// TIA Portal project "Inteligenta_szklarnia" (V15.1) (continued)
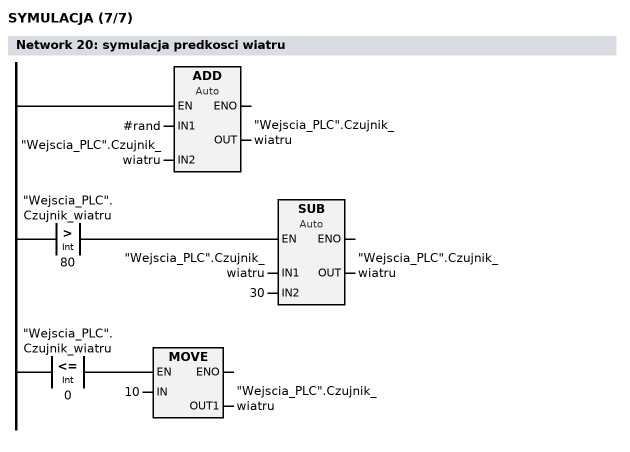
   RUNG wire#powerrail
      Add(in1 := #rand, in2 := "Wejscia_PLC".Czujnik_wiatru, out => "Wejscia_PLC".Czujnik_wiatru)
   END_RUNG
   RUNG wire#powerrail
      { S7_Templates := "SrcType := Int" } GT_Contact(in1 := "Wejscia_PLC".Czujnik_wiatru, in2 := 80)
      Sub(in1 := "Wejscia_PLC".Czujnik_wiatru, in2 := 30, out => "Wejscia_PLC".Czujnik_wiatru)
   END_RUNG
   RUNG wire#powerrail
      { S7_Templates := "SrcType := Int" } LE_Contact(in1 := "Wejscia_PLC".Czujnik_wiatru, in2 := 0)
      Move(in := 10, out1 => "Wejscia_PLC".Czujnik_wiatru)
   END_RUNG
   // the same network as SCL:
   "Wejscia_PLC".Czujnik_wiatru := #rand + "Wejscia_PLC".Czujnik_wiatru;
   IF "Wejscia_PLC".Czujnik_wiatru > 80 THEN
       "Wejscia_PLC".Czujnik_wiatru := "Wejscia_PLC".Czujnik_wiatru - 30;
   END_IF;
   IF "Wejscia_PLC".Czujnik_wiatru <= 0 THEN "Wejscia_PLC".Czujnik_wiatru := 10; END_IF;
END_REGION
END_FUNCTION

ORGANIZATION_BLOCK "Main"   // OB1, LAD, ProgramCycle
TITLE = "Main Program Sweep (Cycle)"
{ S7_Optimized_Access := 'TRUE' }
VERSION : 0.1
   VAR_INPUT
      Initial_Call : Bool;   // Initial call of this OB
      Remanence : Bool;   // =True, if remanent data are available
   END_VAR
   VAR_TEMP   // added for the SCL form of the ladder/FBD networks
      _w1 : Bool;
   END_VAR
BEGIN

REGION Network 1
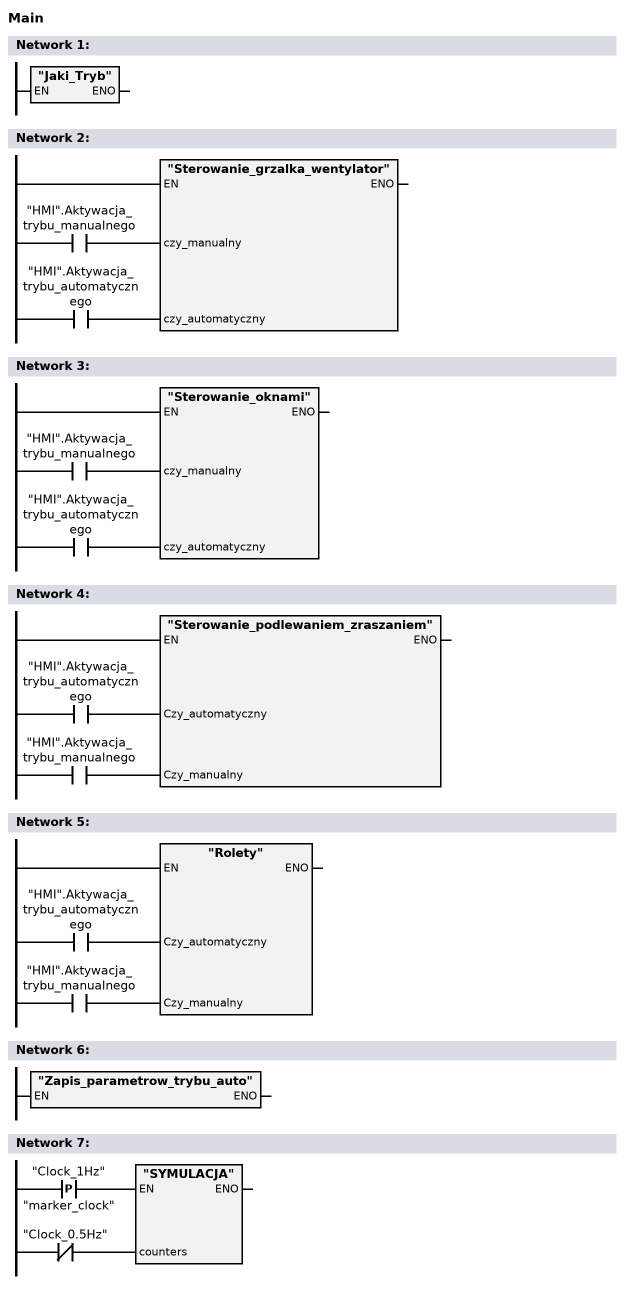
   RUNG wire#powerrail
      "Jaki_Tryb"()
   END_RUNG
   // the same network as SCL:
   "Jaki_Tryb"();
END_REGION

REGION Network 2
   RUNG wire#powerrail
      "Sterowanie_grzalka_wentylator"(czy_manualny := wire#w1, czy_automatyczny := wire#w2)
   END_RUNG
   RUNG wire#powerrail
      Contact( "HMI".Aktywacja_trybu_manualnego )
   END_RUNG wire#w1
   RUNG wire#powerrail
      Contact( "HMI".Aktywacja_trybu_automatycznego )
   END_RUNG wire#w2
   // the same network as SCL:
   "Sterowanie_grzalka_wentylator"(czy_manualny := "HMI".Aktywacja_trybu_manualnego,
                           czy_automatyczny := "HMI".Aktywacja_trybu_automatycznego);
END_REGION

REGION Network 3
   RUNG wire#powerrail
      "Sterowanie_oknami"(czy_manualny := wire#w1, czy_automatyczny := wire#w2)
   END_RUNG
   RUNG wire#powerrail
      Contact( "HMI".Aktywacja_trybu_manualnego )
   END_RUNG wire#w1
   RUNG wire#powerrail
      Contact( "HMI".Aktywacja_trybu_automatycznego )
   END_RUNG wire#w2
   // the same network as SCL:
   "Sterowanie_oknami"(czy_manualny := "HMI".Aktywacja_trybu_manualnego,
                       czy_automatyczny := "HMI".Aktywacja_trybu_automatycznego);
END_REGION

REGION Network 4
   RUNG wire#powerrail
      "Sterowanie_podlewaniem_zraszaniem"(Czy_automatyczny := wire#w1, Czy_manualny := wire#w2)
   END_RUNG
   RUNG wire#powerrail
      Contact( "HMI".Aktywacja_trybu_automatycznego )
   END_RUNG wire#w1
   RUNG wire#powerrail
      Contact( "HMI".Aktywacja_trybu_manualnego )
   END_RUNG wire#w2
   // the same network as SCL:
   "Sterowanie_podlewaniem_zraszaniem"(Czy_automatyczny := "HMI".Aktywacja_trybu_automatycznego,
                           Czy_manualny := "HMI".Aktywacja_trybu_manualnego);
END_REGION

REGION Network 5
   RUNG wire#powerrail
      "Rolety"(Czy_automatyczny := wire#w1, Czy_manualny := wire#w2)
   END_RUNG
   RUNG wire#powerrail
      Contact( "HMI".Aktywacja_trybu_automatycznego )
   END_RUNG wire#w1
   RUNG wire#powerrail
      Contact( "HMI".Aktywacja_trybu_manualnego )
   END_RUNG wire#w2
   // the same network as SCL:
   "Rolety"(Czy_automatyczny := "HMI".Aktywacja_trybu_automatycznego,
            Czy_manualny := "HMI".Aktywacja_trybu_manualnego);
END_REGION

REGION Network 6
   RUNG wire#powerrail
      "Zapis_parametrow_trybu_auto"()
   END_RUNG
   // the same network as SCL:
   "Zapis_parametrow_trybu_auto"();
END_REGION

REGION Network 7
   RUNG wire#powerrail
      P_Contact(operand := "Clock_1Hz", bit := "marker_clock")
      "SYMULACJA"(counters := wire#w1)
   END_RUNG
   RUNG wire#powerrail
      I_Contact( "Clock_0.5Hz" )
   END_RUNG wire#w1
   // the same network as SCL:
   #_w1 := "Clock_1Hz" AND NOT "marker_clock";   // rising edge of "Clock_1Hz"
   "marker_clock" := "Clock_1Hz";
   IF #_w1 THEN "SYMULACJA"(counters := NOT "Clock_0.5Hz"); END_IF;
END_REGION
END_ORGANIZATION_BLOCK

// folder: Archiwizacja_parametrow

FUNCTION "Archiwizacja_parametrow" : Void   // FC2, LAD
{ S7_Optimized_Access := 'TRUE' }
VERSION : 0.1
// Zapis parametrów do bloku DB odbywa się co pół godziny. Po uruchomieniu sterownika pierwszy zapis nie odbywa się od razu, aby wykres nie przedstawiał parametrów, które nie były jeszcze regulowane. Oczytane watosci zapisywane są w tablicach w bloku DB.
   VAR CONSTANT
      iterator : Int := 0;
   END_VAR
   VAR_TEMP   // added for the SCL form of the ladder/FBD networks
      _w1 : Bool;
   END_VAR
BEGIN

REGION Network 1
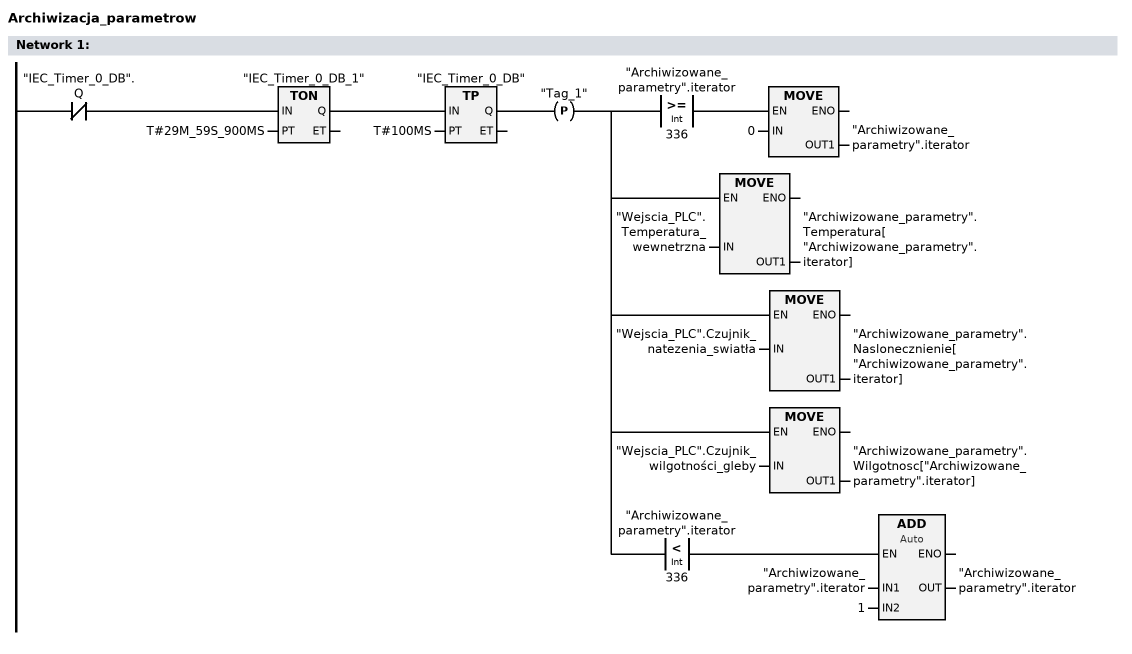
   "IEC_Timer_0_DB_1".TON(IN := NOT "IEC_Timer_0_DB".Q, PT := T#29M_59S_900MS);
   "IEC_Timer_0_DB".TP(IN := "IEC_Timer_0_DB_1".Q, PT := T#100MS);
   #_w1 := "IEC_Timer_0_DB".Q AND NOT "Tag_1";   // rising edge
   "Tag_1" := "IEC_Timer_0_DB".Q;
   IF #_w1 AND ("Archiwizowane_parametry".iterator >= 336) THEN
       "Archiwizowane_parametry".iterator := 0;
   END_IF;
   IF #_w1 THEN
       "Archiwizowane_parametry".Temperatura["Archiwizowane_parametry".iterator] := "Wejscia_PLC".Temperatura_wewnetrzna;
       "Archiwizowane_parametry".Naslonecznienie["Archiwizowane_parametry".iterator] := "Wejscia_PLC".Czujnik_natezenia_swiatła;
       "Archiwizowane_parametry".Wilgotnosc["Archiwizowane_parametry".iterator] := "Wejscia_PLC".Czujnik_wilgotności_gleby;
   END_IF;
   IF #_w1 AND ("Archiwizowane_parametry".iterator < 336) THEN
       "Archiwizowane_parametry".iterator := "Archiwizowane_parametry".iterator + 1;
   END_IF;
END_REGION
END_FUNCTION

// folder: LGF/4 Math operations

FUNCTION "LGF_RandomRange_Real" : Real   // FC10014, SCL
TITLE = LGF_RandomRange_Real
{ S7_Optimized_Access := 'TRUE' }
AUTHOR : Siemens_Digital_Industries
FAMILY : LGF
NAME : LGF_RandomRange_Real
// This function generates random numbers in defined limits (Datatype Real)
   VAR_INPUT
      minValue : Real;   // minimal Value random can reach / Minimum value of the range of the random number
      maxValue : Real;   // maximal Value random can reach / Maximum value of the range of the random number
   END_VAR
   VAR_OUTPUT
      error : Bool;   // Error if true
      status : Word;   // Status of the function
      subfunctionStatus : Word;   // Status or return value of called FB's, FCs and system blocks
   END_VAR
   VAR_TEMP
      tempTime : DTL;   // System time
      tempNanoSecondInDWord : DWord;   // UDINT converted to DWORD for access to individual bytes
      tempTimeStatus : Word;   // Status of the instruction RD_SYS_T
      tempRandomValue : DWord;   // Random-start-value
      tempNormReal : Real;   // normalized value
   END_VAR
   // Ret_Val : Returns random Real number in predefined range
   VAR CONSTANT
      ZERO : Real := 0.0;   // Zero value in case of error
      MAX_UDINT : UDInt := 4294967295;   // Maximum UDINT value
      SUB_STATUS_NO_ERROR : Word := 16#0000;   // Status: sub function call ends without error
      STATUS_FINISHED_NO_ERROR : Word := 16#0000;   // Status: Execution finished without errors
      ERR_MAX_LESS_MIN : Word := 16#8200;   // Error: The maximum limit number is smaller than the minimum limit number
      ERR_RD_SYS_T : Word := 16#8600;   // Error: System function Read system time returned an error
   END_VAR
BEGIN
   REGION Block info header
     //=============================================================================
     // SIEMENS AG / (c)Copyright 2017
     //-----------------------------------------------------------------------------
     // Title:            LGF_RandomRange_Real
     // Comment/Function: This function generates random numbers in defined limits (Datatype Real)
     // Library/Family:   LGF(Library General Functions)
     // Author:           Siemens Digital Industry Support
     // Tested with:      S7-PLCSIM Advanced V2.0 SP1
     // Engineering:      TIA Portal V15 Update 2
     // Restrictions:     ENO disabled - error handling done by error and status
     // Requirements:     PLC (S7-1200 / S7-1500)
     //-------------------------------------------------------------------------------
     // Change log table:
     // Version  | Date       | Expert in charge       | Changes applied
     //----------|------------|------------------------|------------------------------
     // 01.00.00 19.08.2015  Siemens Industry Online Support
     //                      First released version
     // 01.00.01 02.01.2017  Siemens Industry Online Support
     //                      Upgrade: TIA Portal V14 Update 1
     // 01.00.02 02.03.2017  Siemens Industry Online Support
     //                      Bugfix: FC number
     // 01.00.03 17.08.2018  Siemens Industry Online Support
     //                      Upgrade: TIA V15 Update 2
     // 01.00.04 23.11.2018  Siemens Industry Online Support
     //                      Upgrade: TIA V15.1
     // 01.01.00 13.11.2019  Siemens Industry Presales Support
     //                      Renamed from "LGF_RandomReal" to "LGF_RandomRange_Real"
     //                      Regions, commens and costants are added
     // 03.00.00 23.04.2020  Siemens Industry Support
     //                      Set version to V3.0.0, harmonize the version of the whole library
     //=============================================================================
   END_REGION

   REGION Validation
     // Check if the maximal Value is less than the minimal value
     IF (#minValue > #maxValue) THEN
       #error := true;
       #status := #ERR_MAX_LESS_MIN;
       #subfunctionStatus := #SUB_STATUS_NO_ERROR;
       #LGF_RandomRange_Real := #ZERO;
       RETURN;
     END_IF;

     // Read system time
     #tempTimeStatus := INT_TO_WORD(RD_SYS_T(#tempTime));

     // Check return variable for error
     IF (#tempTimeStatus <> #SUB_STATUS_NO_ERROR) THEN
       #error := true;
       #status := #ERR_RD_SYS_T;
       #subfunctionStatus := #tempTimeStatus;
       #LGF_RandomRange_Real := #ZERO;
       RETURN;
     END_IF;
   END_REGION

   REGION Calculating random number
     // Converting to double word so individual bytes can be addressed
     #tempNanoSecondInDWord := UDINT_TO_DWORD(#tempTime.NANOSECOND);

     // Calculate a random-start-value depending on the time
     #tempRandomValue.%B3 := #tempNanoSecondInDWord.%B0;
     #tempRandomValue.%B2 := #tempNanoSecondInDWord.%B1;
     #tempRandomValue.%B1 := #tempNanoSecondInDWord.%B2;
     #tempRandomValue.%B0 := #tempNanoSecondInDWord.%B3;

     // Norm the calculated random number: 0.0 <= #tempNormReal <= 1.0
     #tempNormReal := UDINT_TO_REAL(DWORD_TO_UDINT(#tempRandomValue)) / UDINT_TO_REAL(#MAX_UDINT);

     // Scale the tempNormReal to be in the range of maxValue and minValue
     #LGF_RandomRange_Real := ((#tempNormReal * (#maxValue - #minValue) + (#minValue)));

     #error := false;
     #status := #STATUS_FINISHED_NO_ERROR;
     #subfunctionStatus := #SUB_STATUS_NO_ERROR;
     // ENO mechanism is not used
     ENO := TRUE;
   END_REGION
END_FUNCTION

(* ===== HMI "HMI_RT_3" =====
system functions are stored by id; their names below are inferred from use
connection "HMI_Connection_4": ETHERNET, SMART_S7_1200_OMS

HMI tags "Default tag table"
   "Tag_ScreenNumber" : UInt, internal

HMI tags "wyjsciaPLC"
   "Alarm_ostrzegwaczy" : Bool = PLC Alarm_ostrzegwaczy AT %Q0.5, 100 ms
   "Grzałka" : Bool = PLC Grzałka AT %Q0.0, 100 ms
   "Pompa_wodna" : Bool = PLC Pompa_wodna AT %Q0.2, 100 ms
   "Rolety_otwieranie" : Bool = PLC Rolety_otwieranie AT %Q0.3, 100 ms
   "Rolety_zamykanie" : Bool = PLC Rolety_zamykanie AT %Q0.4, 100 ms
   "Siłownik_okien_otwieranie" : Bool = PLC Siłownik_okien_otwieranie AT %Q0.6, 100 ms
   "Siłownik_okien_zamykanie" : Bool = PLC Siłownik_okien_zamykanie AT %Q0.7, 100 ms
   "Wentylator" : Bool = PLC Wentylator AT %Q0.1, 100 ms
   "Tag_ScreenNumber(1)" : DInt = PLC Tag_ScreenNumber AT %MD0, 500 ms
   "Parametry_Czujnik_światła" : Int = PLC Parametry.Czujnik_światła, 500 ms
   "Parametry_temeratura" : Real = PLC Parametry.temeratura, 500 ms
   "Parametry_Czujnik_wiatru" : Int = PLC Parametry.Czujnik_wiatru, 500 ms
   "Parametry_Wilgotność_powietrza" : Int = PLC Parametry.Wilgotność_powietrza, 500 ms
   "Parametry_czujnik_CO2" : Int = PLC Parametry.czujnik_CO2, 500 ms
   "Parametry_Wilgotność_gleby" : Int = PLC Parametry.Wilgotność_gleby, 500 ms
   "Wejscia_HMI_Temperatura" : Real = PLC Wejscia_HMI.Temperatura, 500 ms
   "Parametry_stopien_zasloniecia_rolet" : Int = PLC Parametry.stopien_zasloniecia_rolet, 1 s
   "Wejscia_HMI_Zaciemnienie" : Int = PLC Wejscia_HMI.Zaciemnienie, 1 s
   "Receptury_nazwa{0}" : String[254] = PLC Receptury.nazwa[0], 1 s
   "Receptury_nazwa{1}" : String[254] = PLC Receptury.nazwa[1], 1 s
   "Receptury_nazwa{2}" : String[254] = PLC Receptury.nazwa[2], 1 s
   "Receptury_nazwa{3}" : String[254] = PLC Receptury.nazwa[3], 1 s
   "Receptury_nazwa{4}" : String[254] = PLC Receptury.nazwa[4], 1 s
   "Receptury_nazwa{5}" : String[254] = PLC Receptury.nazwa[5], 1 s
   "naslonecznienie_man" : Int = PLC Wejscia_HMI.naslonecznienie_manual, 1 s

HMI tags "USTAWIENIA_HMI"
   "temperatura_ustawiona_man" : Real, internal
   "stopien_otwarcia_okien_man" : Real, internal
   "wilgotnosc_powietrza_man" : Real, internal
   "wilgotnosc_gleby_man" : Real, internal
   "nazwa_receptury" : WString[10], internal
   "system_okien" : Bool, internal
   "AlwaysTRUE" : Bool = PLC AlwaysTRUE AT %M1.2, 1 s

screen "Root screen" 800x480, template "Template_1"
   on GenerateScreen: SetTag("Tag_ScreenNumber", 1)
   Button "Button_3" at 10,270 size 300x90; TextOff 'ZAPISZ NOWĄ RECEPTURĘ'
      on Click: ActivateScreen("zapisz_recepture", 0)
   Button "Button_1" at 10,170 size 300x90; TextOff 'TRYB MANUALNY'
      on Click: ActivateScreen("tryb_manualny", 0)
   Button "Button_2" at 10,70 size 301x90; TextOff 'TRYB AUTOMATYCZNY'
      on Click: ActivateScreen("tryb_automatyczny", 0)
   TextField "Text field_2" at 32,2 size 738x63; Text 'AUTOMATYCZNA SZKLARNIA'
   GraphicView "Graphic view_1" at 370,70 size 392x338; Picture "garden-tools-graphic-clipart-design-free-png"
   Button "Button_4" at 10,370 size 301x90; TextOff 'WYBIERZ RECEPTURĘ'
      on Click: ActivateScreen("wybierz_recepture", 0)
   TextField "Text field_1" at 117,454 size 235x26; Text 'Tego przycisku w symulacji nie widac ale nie chciałem uswac jakby jednak był potrzebny xd'
      Visibility <- "AlwaysTRUE"

screen "zapisz_recepture" 800x480
   TextField "Text field_1" at 282,4 size 253x34; Text 'ZAPISZ RECEPTURE / ZAPISZ RECEPTURĘ'
   Button "Button_1" at 750,0 size 50x50; TextOff 'WRÓĆ'; PictureOff "Back_arrow"
      on Click: function_efd93a16()
   Button "Button_2" at 406,414 size 371x53; TextOff 'ZATWIERDŹ'
      on Click: ActivateScreen("praca", 0)
   Bar "Bar_1" at 17,122 size 70x314; MinimumValue 0; MaximumValue 45
      ProcessValue <- "temperatura_ustawiona_man"
   TextField "Text field_2" at 30,64 size 132x23; Text 'TEMPERATURA'
   Bar "Bar_2" at 223,133 size 54x113; MinimumValue 0; MaximumValue 100
      ProcessValue <- "wilgotnosc_powietrza_man"
   TextField "Text field_3" at 231,45 size 122x42; Text 'WOLGOTNOŚĆ POWIETRZA'
   Button "Button_3" at 115,140 size 73x45; TextOff '+ / +0.5 °C'
      on Press: function_dd21b452("temperatura_ustawiona_man", 0.5)
   Button "Button_7" at 115,201 size 73x45; TextOff '- / -0.5 °C'
      on Press: function_b9b71300("temperatura_ustawiona_man", 0.5)
   TextField "Text field_8" at 93,325 size 109x42; Text 'ustawiona wartość USTAWIONA'
   IOField "I/O field_2" at 106,365 size 62x40; FormatPattern 99.9
      ProcessValue <- "temperatura_ustawiona_man"
   TextField "Text field_11" at 156,367 size 37x37; Text '°C'
   Bar "Bar_4" at 225,346 size 57x127; MinimumValue 0; MaximumValue 100
      ProcessValue <- "wilgotnosc_gleby_man"
   TextField "Text field_10" at 229,254 size 122x42; Text 'WOLGOTNOŚĆ GLEBY'
   Button "Button_8" at 230,300 size 40x40; TextOff '+'
      on Click: function_dd21b452("wilgotnosc_gleby_man", 2)
   Button "Button_9" at 318,300 size 40x40; TextOff '-'
      on Click: function_b9b71300("wilgotnosc_gleby_man", 2)
   IOField "I/O field_5" at 291,401 size 62x40; FormatPattern 999
      ProcessValue <- "wilgotnosc_gleby_man"
   TextField "Text field_12" at 285,384 size 83x20; Text 'USTAWIONA'
   TextField "Text field_14" at 338,404 size 30x29; Text '%'
   Button "Button_10" at 223,87 size 40x40; TextOff '+'
      on Click: function_dd21b452("wilgotnosc_powietrza_man", 5)
   Button "Button_11" at 311,87 size 40x40; TextOff '-'
      on Click: function_b9b71300("wilgotnosc_powietrza_man", 5)
   IOField "I/O field_4" at 291,180 size 62x40; FormatPattern 999
      ProcessValue <- "wilgotnosc_powietrza_man"
   TextField "Text field_16" at 288,167 size 83x20; Text 'USTAWIONA'
   TextField "Text field_18" at 342,184 size 30x29; Text '%'
   Button "Button_14" at 3,1 size 43x43; TextOff 'DOM'; PictureOff "home_1"
      on Click: ActivateScreen("Root screen", 0)
   TextField "Text field_4" at 529,47 size 128x23; Text 'SYSTEM OKIEN'
   Switch "Switch_1" at 503,78 size 185x35; TextOn 'ON'; CaptionText 'Switch'; TextOff 'OFF'
      ProcessValue <- "system_okien"
   IOField "I/O field_1" at 426,311 size 328x81; FormatPattern ????????????????????
      ProcessValue <- "nazwa_receptury"
   TextField "Text field_7" at 406,273 size 380x37; Text 'WPISZ NAZWĘ RECEPTURY'
   GraphicView "Graphic view_1" at 385,338 size 36x30; Picture "Graphic_4"
   GraphicView "Graphic view_2" at 753,338 size 36x30; Picture "Graphic_5"
   TextField "Text field_9" at 387,146 size 161x61; Text 'STOPIEŃ OTWARCIA OKIEN ŚREDNIE NASŁONECZNIENIE'
   Bar "Bar_6" at 404,213 size 373x52; MinimumValue 0; MaximumValue 1500
      ProcessValue <- "naslonecznienie_man"
   Button "Button_4" at 697,145 size 80x50; TextOff '+ / -'
      on Click: function_b9b71300("naslonecznienie_man", 5)
   Button "Button_5" at 589,145 size 80x50; TextOff '- / +'
      on Press: function_dd21b452("naslonecznienie_man", 5)

screen "tryb_manualny" 800x480
   Button "Button_2" at 355,415 size 431x53; TextOff 'ZATWIERDŹ'
      on Click: ActivateScreen("praca", 0)
   TextField "Text field_1" at 282,4 size 223x34; Text 'TRYB MANUALNY'
   Bar "Bar_1" at 181,300 size 60x172; MinimumValue 0; MaximumValue 45
      ProcessValue <- "Parametry_temeratura"
   TextField "Text field_2" at 188,267 size 132x23; Text 'TEMPERATURA'
   Bar "Bar_2" at 181,93 size 60x160; MinimumValue 0; MaximumValue 100
      ProcessValue <- "Parametry_Wilgotność_powietrza"
   TextField "Text field_3" at 198,45 size 122x42; Text 'WOLGOTNOŚĆ POWIETRZA WILGOTNOŚĆ POWIETRZA'
   Bar "Bar_3" at 576,166 size 170x52; MinimumValue 0
      ProcessValue <- "stopien_otwarcia_okien_man"
   TextField "Text field_4" at 576,43 size 186x61; Text 'STOPIEŃ OTWARCIA OKIEN STOPIEŃ OTWARCIA OKIEN'
   IOField "I/O field_1" at 244,368 size 95x40; FormatPattern 99.9
      ProcessValue <- "Wejscia_HMI_Temperatura"
   Bar "Bar_4" at 8,93 size 60x160; MinimumValue 0; MaximumValue 100
      ProcessValue <- "Parametry_Wilgotność_gleby"
   Button "Button_4" at 406,253 size 80x60; TextOff 'PODLEWANIE'
      on Click: InvertBit("Pompa_wodna")
   Button "Button_5" at 536,253 size 80x60; TextOff 'GRZANIE'
      on Click: InvertBit("Grzałka")
   Button "Button_6" at 666,253 size 80x60; TextOff 'WENTYLACJA'
      on Click: InvertBit("Wentylator")
   GraphicView "Graphic view_1" at 675,320 size 60x60; Picture "fan_4829316"
      Visibility <- "Wentylator"
   GraphicView "Graphic view_6" at 545,320 size 60x60; Picture "heater_4463010"
      Visibility <- "Grzałka"
   GraphicView "Graphic view_7" at 415,320 size 60x60; Picture "irrigation_18631825"
      Visibility <- "Pompa_wodna"
   GraphicView "Graphic view_9" at 676,320 size 60x60; Picture "fan_off"
      Visibility <- "Wentylator"
   GraphicView "Graphic view_10" at 546,320 size 60x60; Picture "heater_off"
      Visibility <- "Grzałka"
   GraphicView "Graphic view_11" at 415,320 size 60x60; Picture "irrigation_off"
      Visibility <- "Pompa_wodna"
   TextField "Text field_10" at 18,45 size 122x42; Text 'WOLGOTNOŚĆ GLEBY WILGOTNOŚĆ GLEBY'
   IOField "I/O field_3" at 760,171 size 33x36; FormatPattern 9
      ProcessValue <- "stopien_otwarcia_okien_man"
   IOField "I/O field_6" at 70,148 size 62x40; FormatPattern 999
      ProcessValue <- "Parametry_Wilgotność_gleby"
   TextField "Text field_15" at 115,152 size 35x34; Text '%'
   IOField "I/O field_7" at 252,151 size 62x40; FormatPattern 999
      ProcessValue <- "Parametry_Wilgotność_powietrza"
   TextField "Text field_19" at 294,154 size 35x34; Text '%'
   Button "Button_12" at 576,99 size 50x50; TextOff '+'
      on Click: function_dd21b452("stopien_otwarcia_okien_man", 1)
   Button "Button_13" at 696,98 size 50x50; TextOff '-'
      on Click: function_b9b71300("stopien_otwarcia_okien_man", 1)
   Button "Button_14" at 3,1 size 43x43; TextOff 'DOM'; PictureOff "home_1"
      on Click: ActivateScreen("Root screen", 0)
   Button "Button_1" at 750,0 size 50x50; TextOff 'Text'; PictureOff "Back_arrow"
      on Click: function_efd93a16()
   TextField "Text field_9" at 293,369 size 35x34; Text '°C'
   Circle "Circle_1" at 386,336 size 25x25
      Visibility <- "Pompa_wodna"
   Circle "Circle_4" at 386,336 size 25x25
      Visibility <- "Pompa_wodna"
   Circle "Circle_2" at 511,336 size 25x25
      Visibility <- "Grzałka"
   Circle "Circle_5" at 511,336 size 25x25
      Visibility <- "Grzałka"
   Circle "Circle_3" at 639,336 size 25x25
      Visibility <- "Wentylator"
   Circle "Circle_6" at 639,336 size 25x25
      Visibility <- "Wentylator"
   Bar "Bar_5" at 10,300 size 60x172; MinimumValue 0; MaximumValue 1500
      ProcessValue <- "Parametry_Czujnik_światła"
   TextField "Text field_5" at 3,268 size 161x23; Text 'TEMPERATURA / NASŁONECZNIENIE'
   IOField "I/O field_2" at 70,368 size 95x40; FormatPattern 9999
      ProcessValue <- "Parametry_Czujnik_światła"
   TextField "Text field_6" at 127,356 size 35x64; Text '°C W m'
   TextField "Text field_7" at 152,391 size 31x17; Text '2'
   TextField "Text field_8" at 348,43 size 206x61; Text 'STOPIEŃ OTWARCIA OKIEN STOPIEŃ ZASŁONIENIA ROLET'
   Bar "Bar_6" at 366,166 size 170x52; MinimumValue 0; MaximumValue 100
      ProcessValue <- "naslonecznienie_man"
   Button "Button_3" at 456,98 size 80x50; TextOff '+ / ODSŁOŃ'
      on Click: function_b9b71300("naslonecznienie_man", 5)
   Button "Button_7" at 366,98 size 80x50; TextOff '- / ZASŁOŃ'
      on Press: function_dd21b452("naslonecznienie_man", 5)

screen "wybierz_recepture" 800x480
   TextField "Text field_2" at 257,4 size 280x34; Text 'WYBIERZ RECEPTURE / WYBIERZ RECEPTURĘ'
   Button "Button_1" at 750,0 size 50x50; TextOff 'WRÓĆ'; PictureOff "Back_arrow"
      on Click: function_efd93a16()
   Button "Button_14" at 3,1 size 43x43; TextOff 'DOM'; PictureOff "home_1"
      on Click: ActivateScreen("Root screen", 0)
   TextField "Text field_1" at 18,52 size 23x39; Text '1'
   TextField "Text field_3" at 18,108 size 23x39; Text '2'
   TextField "Text field_4" at 18,169 size 23x39; Text '3'
   TextField "Text field_5" at 18,231 size 23x39; Text '4'
   TextField "Text field_6" at 18,290 size 23x39; Text '5'
   TextField "Text field_7" at 18,351 size 23x39; Text '6'
   Button "Button_2" at 13,415 size 775x55; TextOff '-ZATWIERDŹ-'
      on Click: ActivateScreen("praca", 0)
   Button "Button_3" at 720,68 size 60x60; TextOff 'Text'; PictureOff "Double_up_arrow"
   Button "Button_4" at 720,162 size 60x60; TextOff 'Text'; PictureOff "Double_down_arrow"
   Button "Button_5" at 708,326 size 83x64; TextOff 'USUŃ'
   IOField "I/O field_1" at 90,58 size 243x32; FormatPattern ????????????????????
      ProcessValue <- "Receptury_nazwa{0}"
   IOField "I/O field_2" at 90,115 size 241x32; FormatPattern ????????????????????
      ProcessValue <- "Receptury_nazwa{1}"
   IOField "I/O field_3" at 90,176 size 267x32; FormatPattern ????????????????????
      ProcessValue <- "Receptury_nazwa{2}"
   IOField "I/O field_4" at 90,238 size 264x32; FormatPattern ????????????????????
      ProcessValue <- "Receptury_nazwa{3}"
   IOField "I/O field_5" at 90,294 size 230x32; FormatPattern ????????????????????
      ProcessValue <- "Receptury_nazwa{4}"
   IOField "I/O field_6" at 90,358 size 506x32; FormatPattern ????????????????????
      ProcessValue <- "Receptury_nazwa{5}"

screen "praca" 800x480
   GraphicView "Graphic view_2" at 28,217 size 100x100; Picture "Thermometer_icon"
   GraphicView "Graphic view_4" at 276,362 size 100x100; Picture "soil-sensor_11298794"
   GraphicView "Graphic view_3" at 28,74 size 100x100; Picture "sensor_4212513"
   GraphicView "Graphic view_5" at 276,75 size 100x100; Picture "sensor_4212519"
   GraphicView "Graphic view_1" at 559,362 size 100x100; Picture "fan_4829316"
      Visibility <- "Wentylator"
   GraphicView "Graphic view_6" at 560,217 size 100x100; Picture "heater_4463010"
      Visibility <- "Grzałka"
   GraphicView "Graphic view_7" at 560,75 size 100x100; Picture "irrigation_18631825"
      Visibility <- "Pompa_wodna"
   GraphicView "Graphic view_8" at 28,362 size 100x100; Picture "anemometer_1113716"
   GraphicView "Graphic view_9" at 560,362 size 100x100; Picture "fan_off"
      Visibility <- "Wentylator"
   GraphicView "Graphic view_10" at 561,217 size 100x100; Picture "heater_off"
      Visibility <- "Grzałka"
   GraphicView "Graphic view_11" at 561,75 size 100x100; Picture "irrigation_off"
      Visibility <- "Pompa_wodna"
   GraphicView "Graphic view_12" at 276,217 size 100x100; Picture "sensor_2828470"
   TextField "Text field_1" at 54,52 size 204x23; Text 'INSOLATION / NASŁONECZNIENIE / SONNENEINSTRAHLUNG'
   TextField "Text field_2" at 67,194 size 132x23; Text 'TEMPERATURA'
   TextField "Text field_3" at 46,334 size 166x23; Text 'SZYBKOŚĆ WIATRU'
   TextField "Text field_4" at 349,194 size 123x23; Text 'STĘŻENIE CO2'
   TextField "Text field_5" at 294,50 size 223x23; Text 'WILGOTNOŚĆ POWIETRZA'
   TextField "Text field_6" at 321,339 size 175x23; Text 'WILGOTNOŚĆ GLEBY'
   TextField "Text field_7" at 626,46 size 116x23; Text 'PODLEWANIE'
   TextField "Text field_8" at 643,192 size 80x23; Text 'GRZANIE'
   TextField "Text field_9" at 626,330 size 117x23; Text 'WENTYLACJA'
   TextField "Text field_10" at 282,4 size 256x34; Text 'PODGLĄD NA ŻYWO'
   Button "Button_1" at 750,0 size 50x50; TextOff 'WRÓĆ'; PictureOff "Back_arrow"
      on Click: function_efd93a16()
   Button "Button_2" at 3,1 size 43x43; TextOff 'DOM'; PictureOff "home_1"
      on Click: ActivateScreen("Root screen", 0)
   IOField "I/O field_2" at 120,233 size 97x65; FormatPattern 99.99
      ProcessValue <- "Parametry_temeratura"
   IOField "I/O field_3" at 136,383 size 70x65; FormatPattern 999
      ProcessValue <- "Parametry_Czujnik_wiatru"
   IOField "I/O field_5" at 377,235 size 83x65; FormatPattern 9999
      ProcessValue <- "Parametry_czujnik_CO2"
   TextField "Text field_11" at 214,241 size 46x46; Text '°C'
   IOField "I/O field_4" at 406,95 size 69x65; FormatPattern 999
      ProcessValue <- "Parametry_Wilgotność_powietrza"
   IOField "I/O field_6" at 406,384 size 68x65; FormatPattern 999
      ProcessValue <- "Parametry_Wilgotność_gleby"
   TextField "Text field_12" at 472,106 size 47x46; Text '%'
   TextField "Text field_13" at 472,396 size 47x46; Text '%'
   TextField "Text field_14" at 219,90 size 47x72; Text 'W m²'
   IOField "I/O field_1" at 119,109 size 101x32; FormatPattern 99999
      ProcessValue <- "Parametry_Czujnik_światła"
   TextField "Text field_15" at 210,376 size 52x72; Text 'Km h'
   Circle "Circle_1" at 695,101 size 48x48
      Visibility <- "Pompa_wodna"
   Circle "Circle_2" at 695,243 size 48x48
      Visibility <- "Grzałka"
   TextField "Text field_16" at 472,242 size 69x39; Text 'ppm'
   Circle "Circle_4" at 695,101 size 48x48
      Visibility <- "Pompa_wodna"
   Circle "Circle_5" at 695,243 size 48x48
      Visibility <- "Grzałka"
   Circle "Circle_3" at 695,385 size 48x48
      Visibility <- "Wentylator"
   Circle "Circle_6" at 695,385 size 48x48
      Visibility <- "Wentylator"

screen "tryb_automatyczny" 800x480
   IOField "I/O field_1" at 100,354 size 57x40; FormatPattern 99.9
      ProcessValue <- "Wejscia_HMI_Temperatura"
   Button "Button_1" at 750,0 size 50x50; TextOff 'WRÓĆ'; PictureOff "Back_arrow"
      on Click: function_efd93a16()
   Button "Button_2" at 417,418 size 371x53; TextOff 'ZATWIERDŹ'
      on Click: ActivateScreen("praca", 0)
   Bar "Bar_1" at 14,103 size 70x275; MinimumValue 0; MaximumValue 45
      ProcessValue <- "temperatura_ustawiona_man"
   TextField "Text field_2" at 15,60 size 132x23; Text 'TEMPERATURA'
   Bar "Bar_2" at 217,108 size 70x275; MinimumValue 0; MaximumValue 100
      ProcessValue <- "wilgotnosc_powietrza_man"
   TextField "Text field_3" at 205,61 size 122x42; Text 'WOLGOTNOŚĆ POWIETRZA WILGOTNOŚĆ POWIETRZA'
   Button "Button_3" at 90,119 size 75x45; TextOff '+ / +0.5 °C'
      on Press: function_dd21b452("temperatura_ustawiona_man", 0.5)
   Button "Button_7" at 89,177 size 75x45; TextOff '- / -0.5 °C'
      on Press: function_b9b71300("temperatura_ustawiona_man", 0.5)
   IOField "I/O field_2" at 100,276 size 62x40; FormatPattern 99.9
      ProcessValue <- "temperatura_ustawiona_man"
   TextField "Text field_11" at 155,285 size 23x22; Text '°C'
   TextField "Text field_9" at 155,358 size 23x22; Text '°C'
   Bar "Bar_4" at 417,105 size 70x275; MinimumValue 0; MaximumValue 100
      ProcessValue <- "wilgotnosc_gleby_man"
   TextField "Text field_10" at 404,58 size 122x42; Text 'WOLGOTNOŚĆ GLEBY WILGOTNOŚĆ GLEBY'
   Button "Button_8" at 496,125 size 65x40; TextOff '+ / +2%'
      on Click: function_dd21b452("wilgotnosc_gleby_man", 2)
   Button "Button_9" at 497,177 size 65x40; TextOff '- / -2%'
      on Click: function_b9b71300("wilgotnosc_gleby_man", 2)
   IOField "I/O field_5" at 508,276 size 62x40; FormatPattern 999
      ProcessValue <- "wilgotnosc_gleby_man"
   IOField "I/O field_6" at 508,346 size 62x40; FormatPattern 999
      ProcessValue <- "Parametry_Wilgotność_gleby"
   TextField "Text field_12" at 493,264 size 101x22; Text 'USTAWIONA'
   TextField "Text field_13" at 497,335 size 86x22; Text 'AKTUALNA'
   TextField "Text field_14" at 547,285 size 23x22; Text '%'
   TextField "Text field_15" at 547,356 size 23x22; Text '%'
   Button "Button_10" at 298,125 size 65x40; TextOff '+ / +5%'
      on Click: function_dd21b452("wilgotnosc_powietrza_man", 5)
   Button "Button_11" at 298,177 size 65x40; TextOff '- / -5%'
      on Click: function_b9b71300("wilgotnosc_powietrza_man", 5)
   IOField "I/O field_4" at 305,277 size 66x40; FormatPattern 999
      ProcessValue <- "wilgotnosc_powietrza_man"
   IOField "I/O field_7" at 307,349 size 62x40; FormatPattern 999
      ProcessValue <- "Parametry_Wilgotność_powietrza"
   TextField "Text field_16" at 292,264 size 101x22; Text 'USTAWIONA'
   TextField "Text field_17" at 294,335 size 86x22; Text 'AKTUALNA'
   TextField "Text field_18" at 346,286 size 23x22; Text '%'
   TextField "Text field_19" at 346,357 size 23x22; Text '%'
   Button "Button_14" at 3,1 size 43x43; TextOff 'DOM'; PictureOff "home_1"
      on Click: ActivateScreen("Root screen", 0)
   TextField "Text field_4" at 38,424 size 128x23; Text 'SYSTEM OKIEN'
   Switch "Switch_1" at 198,418 size 185x35; TextOn 'ON'; CaptionText 'Switch'; TextOff 'OFF'
      ProcessValue <- "system_okien"
   GraphicView "Graphic view_1" at 150,60 size 40x40; Picture "Thermometer_icon"
   GraphicView "Graphic view_2" at 330,61 size 40x40; Picture "sensor_4212519"
   TextField "Text field_5" at 93,334 size 86x22; Text 'AKTUALNA'
   TextField "Text field_6" at 90,262 size 101x22; Text 'USTAWIONA'
   GraphicView "Graphic view_3" at 526,61 size 40x40; Picture "soil-sensor_11298794"
   TextField "Text field_1" at 250,4 size 288x34; Text 'TRYB AUTOMATYCZNY'
   Bar "Bar_3" at 620,105 size 70x275; MinimumValue 0; MaximumValue 1500
      ProcessValue <- "wilgotnosc_gleby_man"
   TextField "Text field_7" at 604,53 size 161x42; Text 'WOLGOTNOŚĆ GLEBY NASŁONECZNIENIE'
   GraphicView "Graphic view_4" at 725,79 size 40x40; Picture "sensor_4212513"
   Button "Button_4" at 696,125 size 65x40; TextOff '+ +25 W m'
      on Click: function_dd21b452("naslonecznienie_man", 25)
   Button "Button_5" at 697,177 size 65x40; TextOff '- -25 W m'
      on Click: function_b9b71300("naslonecznienie_man", 25)
   IOField "I/O field_3" at 708,276 size 62x40; FormatPattern 999
      ProcessValue <- "naslonecznienie_man"
   TextField "Text field_8" at 693,264 size 101x22; Text 'USTAWIONA'
   IOField "I/O field_8" at 711,347 size 62x40; FormatPattern 999
      ProcessValue <- "Parametry_Czujnik_światła"
   TextField "Text field_20" at 697,335 size 86x22; Text 'AKTUALNA'
   TextField "Text field_21" at 747,285 size 23x22; Text '%'
   TextField "Text field_22" at 747,356 size 23x22; Text '%'
   TextField "Text field_23" at 751,143 size 32x18; Text '2'
   TextField "Text field_24" at 748,196 size 32x18; Text '2'

Template "Template_1" 800x480
   Button "Exit" at 671,429 size 71x50; TextOn 'Exit'; TextOff 'Exit'; PictureOn "ExitRuntime_KTP700_Basic_PN_TR"; PictureOff "ExitRuntime_KTP700_Basic_PN_TR"
      on Release: StopRuntime(0)
   Button "Alarms" at 524,429 size 71x50; TextOn 'Alarms'; TextOff 'Alarms'; PictureOn "AlarmDisplay_KTP700_Basic_PN_TR"; PictureOff "AlarmDisplay_KTP700_Basic_PN_TR"
      on Release: function_ef3f5d25("Alarm window_Unacknowledged", -1)
   Button "Start screen" at 169,429 size 71x50; TextOn 'Start screen'; TextOff 'Start screen'; PictureOn "NavigateHome_KTP700_Basic_PN_TR"; PictureOff "NavigateHome_KTP700_Basic_PN_TR"
      on Release: ActivateScreen("Root screen", 0)
      Visibility <- "AlwaysTRUE"
   Button "Language" at 377,429 size 71x50; TextOn 'Language'; TextOff 'Language'; PictureOn "ToggleLanguage_KTP700_Basic_PN_TR"; PictureOff "ToggleLanguage_KTP700_Basic_PN_TR"
      on Release: function_fb9197e8(-1)
*)

(* ===== HMI "HMI_RT_2" =====
system functions are stored by id; their names below are inferred from use
connection "HMI_Connection_3": ETHERNET, SMART_S7_1200_OMS

HMI tags "Default tag table"
   "Tag_ScreenNumber" : Int = PLC HMI.Numer_ekranu_HMI AT %MD0, 100 ms
   "AlwaysTRUE" : Bool = PLC AlwaysTRUE AT %M1.2, 1 s
   "HMI_Aktywacja_trybu_zapis_Receptur" : Bool = PLC HMI.Aktywacja_trybu_zapis_Receptur, 1 s
   "HMI_Aktywacja_trybu_Receptur" : Bool = PLC HMI.Aktywacja_trybu_Receptur, 1 s
   "HMI_Aktywacja_trybu_automatycznego" : Bool = PLC HMI.Aktywacja_trybu_automatycznego, 1 s
   "Tryb_auto_parametry_Temperatura" : Real = PLC Tryb_auto_parametry.Temperatura, 1 s
   "Tryb_auto_parametry_System_okien" : Bool = PLC Tryb_auto_parametry.System_okien, 1 s
   "Tryb_auto_parametry_Wilgotnosc_gleby" : Int = PLC Tryb_auto_parametry.Wilgotnosc_gleby, 1 s
   "Tryb_auto_parametry_Naslonecznienie" : Int = PLC Tryb_auto_parametry.Naslonecznienie, 1 s
   "Tryb_auto_parametry_Stezenie_co2" : Int = PLC Tryb_auto_parametry.Stezenie_co2, 1 s
   "Tryb_auto_parametry_Wilgotnosc_powietrza" : Int = PLC Tryb_auto_parametry.Wilgotnosc_powietrza, 1 s
   "Pompa_zraszacze" : Bool = PLC Pompa_zraszacze AT %Q0.2, 1 s
   "Pompa_podlewanie" : Bool = PLC Pompa_podlewanie AT %Q1.0, 1 s
   "Grzałka" : Bool = PLC Grzałka AT %Q0.0, 1 s
   "Wentylator" : Bool = PLC Wentylator AT %Q0.1, 1 s
   "HMI_Reset_Trybow" : Bool = PLC HMI.Reset_Trybow, 1 s

HMI tags "Do_PLC"
   "System_okien_auto" : Bool = PLC HMI.System_okien_auto, 500 ms
   "Stopien_zasloniecia_rolet_manual" : Int = PLC HMI.Stopien_zasloniecia_rolet_manual, 100 ms
   "Przycisk_zraszania_manual" : Bool = PLC HMI.Przycisk_zraszacze_manual AT %Q0.2, 100 ms
   "Przycisk_wentylacja_manual" : Bool = PLC HMI.Przycisk_wentylacja_manual AT %Q0.1, 100 ms
   "Przycisk_grzanie_manual" : Bool = PLC HMI.Przycisk_grzanie_manual AT %Q0.0, 100 ms
   "Otwarcie_okien_man" : Bool = PLC HMI.Otwarcie_okien_manual AT %DB1.DBW0, 100 ms
   "Temperatura_auto" : Real = PLC HMI.Temperatura_auto, 500 ms
   "Naslonecznienie_auto" : Int = PLC HMI.Naslonecznienie_auto AT %DB1.DBW0, 500 ms
   "Wilgotnosc_powietrza_auto" : Int = PLC HMI.Wilgotnosc_powietrza_auto AT %DB1.DBW0, 500 ms
   "Wilgotnosc_gleby_auto" : Int = PLC HMI.Wilgotnosc_gleby_auto AT %DB1.DBW0, 500 ms
   "Przycisk_zatwierdz_auto" : Bool = PLC HMI.Przycisk_zatwierdz_auto AT %DB1.DBW0, 100 ms
   "nazwa_receptury" : String[254] = PLC HMI.nazwa_receptury AT %DB1.DBX0.0, 500 ms
   "przycisk_zatwierdz_zapis_receptury" : Bool = PLC HMI.Przycisk_zatwierdz_zapis_receptury AT %DB1.DBX0.0, 500 ms
   "HMI_Przycisk_zatwierdz_wybor_receptury" : Bool = PLC HMI.Przycisk_zatwierdz_wybor_receptury AT %DB1.DBX0.0, 500 ms
   "Przycisk_podlewania_manual" : Bool = PLC HMI.Przycisk_podlewanie_manual AT %Q0.2, 100 ms
   "Poziom_CO2_auto" : Int = PLC HMI.Poziom_CO2_auto AT %DB1.DBX0.0, 1 s

HMI tags "Z_PLC"
   "Czujnik_wilgotności_powietrza" : Int = PLC Wejscia_PLC.Czujnik_wilgotności_powietrza, 500 ms
   "Temperatura_wewnetrzna" : Real = PLC Wejscia_PLC.Temperatura_wewnetrzna, 500 ms
   "Czujnik_natezenia_światła" : Int = PLC Wejscia_PLC.Czujnik_natezenia_swiatła, 500 ms
   "Czujnik_wilgotności_gleby" : Int = PLC Wejscia_PLC.Czujnik_wilgotności_gleby, 500 ms
   "Wewnetrzny_czujnik_CO2" : Int = PLC Wejscia_PLC.Wewnetrzny_czujnik_CO2, 500 ms
   "Czujnik_wiatru" : Int = PLC Wejscia_PLC.Czujnik_wiatru, 500 ms
   "Stopien_zasloniecia_rolet" : Int = PLC Wejscia_PLC.Stopien_zasloniecia_rolet, 1 s
   "Zewnetrzny_czujnik_CO2" : Int = PLC Wejscia_PLC.Zewnetrzny_czujnik_CO2 AT %DB1.DBW0, 1 s
   "Temperatura_zewnetrzna" : Real = PLC Wejscia_PLC.Temperatura_zewnetrzna AT %DB1.DBW0, 1 s

text list "receptury": 0..1 ''

recipe "Receptura_nr1": Temperatura <- "Tryb_auto_parametry_Temperatura", Wilgotność Powietrza <- "Tryb_auto_parametry_Wilgotnosc_powietrza", Wilgotność gleby <- "Tryb_auto_parametry_Wilgotnosc_gleby", System okien <- "Tryb_auto_parametry_System_okien", Stężenie CO2 <- "Tryb_auto_parametry_Stezenie_co2", Nasłonecznienie <- "Tryb_auto_parametry_Naslonecznienie"

screen "Root screen" 800x480, template "Template_1"
   on GenerateScreen: SetTag("Tag_ScreenNumber", 0)
   Button "Button_1" at 9,154 size 300x70; TextOff 'TRYB MANUALNY'
      on Click: ActivateScreen("tryb_manualny", 0)
   Button "Button_2" at 10,70 size 300x70; TextOff 'TRYB AUTOMATYCZNY'
      on Click: ActivateScreen("tryb_automatyczny", 0)
   TextField "Text field_2" at 32,2 size 738x63; Text 'AUTOMATYCZNA SZKLARNIA'
   GraphicView "Graphic view_1" at 370,70 size 392x338; Picture "garden-tools-graphic-clipart-design-free-png"
   Button "Button_5" at 10,237 size 300x70; TextOff 'TRYB RECEPTUR'
      on Click: function_e3503463('\USB_X60.1\record.csv', U 0, 2, 1, N); ActivateScreen("Receptury", 0)
   Button "Button_3" at 10,322 size 300x70; TextOff 'SYMULACJA'
      on Click: ActivateScreen("Symulacja_czujnikow", 0)

